
Template "top_menu" 800x480
   Button "Template_Button_3" at 3,3 size 45x34; TextOff 'Text'
      on Click: function_cf6f4242("GraphX_Slidein_Left", -1)
   Group "Group_2" at 3,3 size 45x34
   Group "Group_3" at 747,1 size 53x34
   GraphicView "Template_Graphic view_1" at 69,0 size 40x38; Picture "344330-200"
   Button "BtnBack" at 67,3 size 45x34; TextOff 'Text'
      on Click: function_efd93a16()
   GraphicView "Template_Graphic view_2" at 130,3 size 35x34; Picture "Artboard_43-512"
   Button "BtnHome" at 127,4 size 45x34; TextOff 'Text'
      on Click: ActivateScreen("Main", 0)
   IOField "Template_I/O field_2" at 638,2 size 46x16; FormatPattern 999; Unit  
   IOField "Template_I/O field_3" at 532,18 size 82x16; FormatPattern 999; Unit  
   TextField "Template_Text field_3" at 490,18 size 40x16; Text 'Errors:'
   IOField "Template_I/O field_1" at 614,18 size 70x16; FormatPattern 999; Unit  
   TextField "Template_Text field_1" at 619,19 size 27x16; Text 'Sim:'
   IOField "Template_I/O field_4" at 532,2 size 106x16; FormatPattern 999; Unit  
   TextField "Template_Text field_4" at 643,1 size 10x16; Text '/'
   TextField "Template_Text field_2" at 483,2 size 45x16; Text 'Alarms:'
   Button "Template_Button_2" at 531,1 size 154x34; TextOff 'Text'
   Switch "Template_Switch_1" at 684,1 size 64x34; CaptionText 'Switch'; TextOff 'Tags OFF'; TextOn 'Tags ON'
   Button "Template_Button_5" at 747,1 size 53x34; TextOff 'Text'
      on Click: function_cf6f4242("GraphX_Slidein_Right", -1)

screen "Main" 800x480, template "top_menu"
   ScreenModuleView "motorValveAnalogIcon_1" at 139,122 size 123x41; Guid_{11997190-91299} 'PT-01'; ScreenModuleType ""
      on Guid_{11997190-75677}: function_efd93a16("Analog1", 50, 50, -1, 0, 1)
   Group "Group" at 265,110 size 32x56
   Group "Group_1" at 56,180 size 42x20
   ScreenModuleView "analogInAndAlarmsIcon_1" at 533,124 size 73x71; Guid_{11997190-95263} 'MV-01'; ScreenModuleType ""
      on Guid_{11997190-75677}: function_efd93a16("Valve1", 30, 30, 1, -1, 1)
   ScreenModuleView "analogInAndAlarmsIcon_2" at 535,284 size 73x71; Guid_{11997190-95263} 'MV-02'; ScreenModuleType ""
      on Guid_{11997190-75677}: function_efd93a16("Valve2", 30, 30, 1, -1, 1)
   Group "Group_2" at 671,178 size 42x20
   Group "Group_3" at 668,342 size 42x20
   ScreenModuleView "motorValveAnalogIcon_2" at 144,282 size 123x41; Guid_{11997190-91299} 'TT-01'; ScreenModuleType ""
      on Guid_{11997190-75677}: function_efd93a16("Analog2", 50, 50, -1, 0, 1)
   TextField "Text field_1" at 269,115 size 24x23; Text 'PT'

PopupScreen "Analog1" 502x247
   ScreenModuleView "analogInAndAlarmsFP_1" at 1,1 size 500x244; ScreenModuleType ""
      Guid_{11997190-61144} <- "example_AI_PT44"
   Button "Button_1" at 429,9 size 57x36; TextOff 'X'
      on Click: function_efd93a16("Analog1", 30, 30, 0, -1, 1)

PopupScreen "Valve1" 502x247
   ScreenModuleView "motorValveFacplate_1" at 2,3 size 499x244; Guid_{11997190-89252} 'Valve 1'; ScreenModuleType ""
      on Guid_{11997190-86333}: function_efd93a16("Valve1", 50, 50, 0, -1, 1)
      Guid_{11997190-61144} <- "example_motorValveAnalog_DB_valve1_hmi"

screen "Alarms" 800x480, template "top_menu"
   AlarmView "Alarm view_1" at 8,42 size 789x432

PopupScreen "Valve2" 502x247
   ScreenModuleView "motorValveFacplate_1" at 2,3 size 499x244; Guid_{11997190-89252} 'Valve_2'; ScreenModuleType ""
      on Guid_{11997190-86333}: function_efd93a16("Valve2", 50, 50, 0, -1, 1)
      Guid_{11997190-61144} <- "example_motorValveAnalog_DB_valve2_hmi"

PopupScreen "Analog2" 502x247
   ScreenModuleView "analogInAndAlarmsFP_1" at 1,1 size 500x244; ScreenModuleType ""
      Guid_{11997190-61144} <- "example_AI_PT44"
   Button "Button_1" at 429,9 size 57x36; TextOff 'X'
      on Click: function_efd93a16("Analog2", 30, 30, 0, -1, 1)

screen "UserMangement" 800x480, template "top_menu"
   UserView "User view_1" at 7,46 size 782x425

screen "Diagnostics" 800x480, template "top_menu"
   SysDiagControl "System diagnostics view_1" at 3,40 size 792x436

screen "Test" 800x480, template "top_menu"
   PLCCodeViewer "PLC code view_1" at 35,84 size 543x266
   S7GraphOverview "GRAPH overview_1" at 159,383 size 424x72

screen "load_balanser" 800x480
   ScreenModuleView "load_balancer_faceplate_1" at 127,122 size 640x320; ScreenModuleType ""

VB script "VBFunction_1"
   'Tip:
   ' 1. Use the <CTRL+SPACE> or <CTRL+I> shortcut to open a list of all objects and functions
   ' 2. Write the code using the HMI Runtime object.
   '  Example: HmiRuntime.Screens("Screen_1").
   ' 3. Use the <CTRL+J> shortcut to create an object reference.
   'Write the code as of this position:
*)

(* ===== HMI "HMI_RT_1" =====
system functions are stored by id; their names below are inferred from use

ScreenModuleEditorView "AnalogInAndAlarmsIcon" 125x43
   Button "value_alarmH" at 104,17 size 16x12; TextOff 'H'
      on Click: SetTag("screen", 3)
      Visibility <- "aiUdt.alarmH.Q"
   Button "value_alarmL" at 104,26 size 16x12; TextOff 'L'
      on Click: SetTag("screen", 3)
      Visibility <- "aiUdt.alarmL.Q"
   Button "value_simulation" at 1,17 size 12x21; TextOff 'SIM'
      Visibility <- "aiUdt.ai.sim"
      Appearance <- "aiUdt.ai.sim"
   IOField "value_value" at 12,17 size 92x21; FormatPattern 99999.99
      ProcessValue <- "aiUdt.ai.Q"
      Appearance <- "aiUdt.ai.Error"
   Button "value_alarmLL" at 104,26 size 16x12; TextOff 'LL'
      on Click: SetTag("screen", 3)
      Visibility <- "aiUdt.alarmLL.Q"
   Button "value_alarmHH" at 104,17 size 16x12; TextOff 'HH'
      on Click: SetTag("screen", 3)
      Visibility <- "aiUdt.alarmHH.Q"
   Button "Button" at 0,1 size 123x40; TextOff 'Text'
   TextField "Text field_1" at 8,-1 size 91x20; Text 'TAG_TAG_TAG'
      Visibility <- "aiUdt.hmi.showTag"

VB script "unitIntervalChange"
   'Tip:
   ' 1. Use the <CTRL+SPACE> or <CTRL+I> shortcut to open a list of all objects and functions
   ' 2. Write the code using the HMI Runtime object. Example: HmiRuntime.Screens("Screen_1").
   ' 3. Use the <CTRL+J> shortcut to create an object reference.
*)

(* ===== HMI "HMI_RT_1" =====
system functions are stored by id; their names below are inferred from use

HMI tags "Default tag table"
   "screen" : Int, internal
   "unitIntervalPerCent" : Real, internal

ScreenModuleEditorView "analogInAndAlarmsFacplate" 500x244
   IOField "I/O field_13" at 228,60 size 66x30; FormatPattern 9999.99
      Visibility <- "screen"
      ProcessValue <- "aiUdt.ai.scaleMin"
   IOField "I/O field_14" at 228,98 size 66x30; FormatPattern 9999.99
      Visibility <- "screen"
      ProcessValue <- "aiUdt.ai.scaleMax"
   IOField "I/O field_15" at 228,140 size 66x30; FormatPattern 9999.99
      Visibility <- "screen"
   IOField "I/O field_16" at 228,178 size 66x30; FormatPattern 9999.99
      Visibility <- "screen"
   IOField "I/O field_17" at 71,59 size 77x30; FormatPattern 99999.99
      Visibility <- "screen"
      ProcessValue <- "aiUdt.ai.Q"
      ObjectEnable <- "aiUdt.ai.sim"
   TextField "Text field_8" at 157,64 size 65x20; Text 'Scale Min:'
      Visibility <- "screen"
   TextField "Text field_9" at 157,101 size 68x20; Text 'Scale Max:'
      Visibility <- "screen"
   TextField "Text field_10" at 157,144 size 46x20; Text 'Factor:'
      Visibility <- "screen"
   TextField "Text field_11" at 157,181 size 33x20; Text 'Bias:'
      Visibility <- "screen"
   TextField "Text field_12" at 7,65 size 42x20; Text 'Value:'
      Visibility <- "screen"
   IOField "I/O field_18" at 407,93 size 69x30; FormatPattern 999; Unit  %
      Visibility <- "screen"
      ProcessValue <- "aiUdt.ai.filterConst"
   TextField "Text field_14" at 308,98 size 73x20; Text 'Error Action'
      Visibility <- "screen"
   IOField "I/O field_19" at 413,58 size 66x30; FormatPattern 999999
      Visibility <- "screen"
      ProcessValue <- "aiUdt.ai.filterConst"
   TextField "Text field_15" at 310,65 size 66x20; Text 'FilterConst'
      Visibility <- "screen"
   TextField "Text field_17" at 6,98 size 55x20; Text 'Simulate'
      Visibility <- "screen"
      Appearance <- "aiUdt.ai.sim"
   TextField "Text field_29" at 307,125 size 78x36; Text 'Force inside scale:'
      Visibility <- "screen"
   IOField "I/O field_23" at 69,136 size 78x30; FormatPattern 999.9; Unit  %
      Visibility <- "screen"
      ProcessValue <- "aiUdt.ai.unitInterval"
   TextField "Text field_30" at 6,143 size 54x20; Text 'Raw val.'
      Visibility <- "screen"
   Button "BtnHelpFilterConst" at 383,61 size 26x24; TextOff '?'
      Visibility <- "screen"
   GraphicView "Graphic view_4" at 32,194 size 32x19; Picture "kisspng-computer-icons-cut-copy-and-paste-copying-clip-a-options-vector-5adbf59dcb7576.1022898415243647018334"
      Visibility <- "screen"
   GraphicView "Graphic view_5" at 83,192 size 24x27; Picture "kisspng-computer-icons-clipboard-cut-copy-and-paste-5ae0cc5c36eb73.140446591524681820225"
      Visibility <- "screen"
   Button "BtnScreenEmpty_7" at 31,188 size 40x31; TextOff 'Text'
      on Click: SetTag(N, 1)
      Visibility <- "screen"
   Button "BtnScreenEmpty_6" at 81,185 size 36x36; TextOff 'Text'
      on Click: SetTag("screen", 201)
      Visibility <- "screen"
   Switch "Switch_2" at 411,134 size 61x30; TextOn 'On'; CaptionText 'Switch'; TextOff 'Off'
      Appearance <- "aiUdt.ai.forceInsideScale"
      ProcessValue <- "aiUdt.ai.forceInsideScale"
      Visibility <- "screen"
   Switch "Switch_1" at 101,96 size 46x25; TextOn 'On'; CaptionText 'Switch'; TextOff 'Off'
      Appearance <- "aiUdt.ai.sim"
      ProcessValue <- "aiUdt.ai.sim"
      Visibility <- "screen"
   Button "BtnScreenEmpty" at 407,179 size 62x40; TextOff '?'
      on Click: SetTag("screen", 300)
      Visibility <- "screen"
   Polyline "Polyline_7" at 428,153 size 25x56
      Visibility <- "screen"
   Rectangle "Rectangle_1" at 98,119 size 75x47
      Visibility <- "screen"
   Polyline "Polyline_1" at 32,127 size 56x25
      Visibility <- "screen"
   TextField "Text field_18" at 23,109 size 47x22; Text 'Raw in'
      Visibility <- "screen"
   TextField "Text field_19" at 103,131 size 64x22; Text 'Run. avg'
      Visibility <- "screen"
   Polyline "Polyline_2" at 189,127 size 56x25
      Visibility <- "screen"
   Rectangle "Rectangle_2" at 253,121 size 73x42
      Visibility <- "screen"
   TextField "Text field_20" at 258,131 size 65x22; Text 'Err check'
      Visibility <- "screen"
   Polyline "Polyline_3" at 125,59 size 25x56
      Visibility <- "screen"
   TextField "Text field_21" at 50,68 size 80x22; Text 'Filter const.'
      Visibility <- "screen"
   Polyline "Polyline_4" at 344,122 size 56x25
      Visibility <- "screen"
   Rectangle "Rectangle_3" at 399,122 size 73x42
      Visibility <- "screen"
   TextField "Text field_22" at 408,131 size 48x22; Text 'Scaling'
      Visibility <- "screen"
   Polyline "Polyline_5" at 420,57 size 25x56
      Visibility <- "screen"
   TextField "Text field_23" at 339,69 size 75x22; Text 'Min & Max'
      Visibility <- "screen"
   Rectangle "Rectangle_4" at 344,197 size 73x42
      Visibility <- "screen"
   TextField "Text field_24" at 151,211 size 59x22; Text 'Simulate'
      Visibility <- "screen"
   Polyline "Polyline_6" at 280,211 size 56x25
      Visibility <- "screen"
   TextField "Text field_25" at 299,206 size 91x22; Text 'Factor & bias'
      Visibility <- "screen"
   Polyline "Polyline_8" at 424,211 size 56x25
      Visibility <- "screen"
   TextField "Text field_26" at 444,195 size 16x22; Text 'Q'
      Visibility <- "screen"
   Button "value_alarmHH" at 18,147 size 36x26; TextOff 'HH'
      on Click: SetTag("screen", 3)
      Visibility <- "screen"
      Appearance <- "aiUdt.alarmHH.Q"
   Button "value_alarmH" at 57,147 size 36x26; TextOff 'H'
      on Click: SetTag("screen", 3)
      Visibility <- "screen"
      Appearance <- "aiUdt.alarmH.Q"
   Button "value_alarmL" at 96,147 size 36x26; TextOff 'L'
      on Click: SetTag("screen", 3)
      Visibility <- "screen"
      Appearance <- "aiUdt.alarmL.Q"
   Button "value_alarmLL" at 135,147 size 36x26; TextOff 'LL'
      on Click: SetTag("screen", 3)
      Visibility <- "screen"
      Appearance <- "aiUdt.alarmLL.Q"
   Button "value_simulation" at 41,184 size 99x35; TextOff 'Simulation'
      Visibility <- "screen"
      Appearance <- "aiUdt.ai.sim"
   Bar "Bar" at 200,63 size 66x171; MinimumValue 0; MaximumValue 100
      MinimumValue <- "aiUdt.ai.scaleMin"
      ProcessValue <- "aiUdt.ai.Q"
      MaximumValue <- "aiUdt.ai.scaleMax"
      Visibility <- "screen"
   IOField "value_value" at 18,74 size 151x42; FormatPattern 99999999; Unit         
      Visibility <- "screen"
      ProcessValue <- "aiUdt.alarmHH.delay"
      Appearance <- "aiUdt.ai.Error"
   GraphicView "Graphic 123" at 33,9 size 40x37; Picture "123-512"
   GraphicView "Graphic gear" at 182,7 size 40x37; Picture "setting-512"
   GraphicView "Graphic alarm" at 109,6 size 40x37; Picture "UI_Glyph_09_-13-512"
   Button "BtnScreenValue" at 22,4 size 57x42; TextOff 'Text'
      on Click: SetTag("screen", 0)
   Button "BtnScreenAlarms" at 97,4 size 57x42; TextOff 'Text'
      on Click: SetTag("screen", 100)
   Button "BtnScreenSetup" at 174,4 size 57x42; TextOff 'Text'
      on Click: SetTag("screen", 200)
   Switch "Switch_10" at 131,197 size 46x27; TextOn 'On'; CaptionText 'Switch'; TextOff 'Off'
      Appearance <- "aiUdt.ai.forceInsideScale"
      Visibility <- "screen"
      ProcessValue <- "aiUdt.alarmLL.autoAck"
   IOField "I/O field_5" at 190,160 size 62x30; FormatPattern 9999.99
      Visibility <- "screen"
      ProcessValue <- "aiUdt.alarmL.lim"
   IOField "I/O field_1" at 190,84 size 62x30; FormatPattern 9999.99
      Visibility <- "screen"
      ProcessValue <- "aiUdt.alarmHH.lim"
   TextField "Text field_1" at 7,91 size 64x20; Text 'Alarm HH:'
      Visibility <- "screen"
   TextField "Text field_2" at 205,63 size 26x17; Text 'Limit'
      Visibility <- "screen"
   TextField "Text field_3" at 268,63 size 56x17; Text 'Delay [ms]'
      Visibility <- "screen"
   IOField "I/O field_2" at 265,84 size 53x30; FormatPattern 99999
      Visibility <- "screen"
      ProcessValue <- "aiUdt.alarmHH.delay"
   IOField "I/O field_3" at 190,121 size 62x30; FormatPattern 9999.99
      Visibility <- "screen"
      ProcessValue <- "aiUdt.alarmH.lim"
   TextField "Text field_4" at 7,125 size 56x20; Text 'Alarm H:'
      Visibility <- "screen"
   IOField "I/O field_4" at 265,121 size 53x30; FormatPattern 99999
      Visibility <- "screen"
      ProcessValue <- "aiUdt.alarmH.delay"
   TextField "Text field_5" at 7,165 size 54x20; Text 'Alarm L:'
      Visibility <- "screen"
   IOField "I/O field_6" at 265,160 size 53x30; FormatPattern 99999
      Visibility <- "screen"
      ProcessValue <- "aiUdt.alarmL.delay"
   IOField "I/O field_7" at 190,197 size 62x30; FormatPattern 9999.99
      Visibility <- "screen"
      ProcessValue <- "aiUdt.alarmLL.lim"
   TextField "Text field_6" at 7,201 size 60x20; Text 'Alarm LL:'
      Visibility <- "screen"
   IOField "I/O field_8" at 265,197 size 53x30; FormatPattern 99999
      Visibility <- "screen"
      ProcessValue <- "aiUdt.alarmLL.delay"
   IOField "I/O field_9" at 331,84 size 67x30; FormatPattern 9999.99
      Visibility <- "screen"
      ProcessValue <- "aiUdt.alarmHH.hyst"
   TextField "Text field_7" at 337,63 size 55x17; Text 'Hysteresis'
      Visibility <- "screen"
   IOField "I/O field_10" at 331,121 size 67x30; FormatPattern 9999.99
      Visibility <- "screen"
      ProcessValue <- "aiUdt.alarmH.hyst"
   IOField "I/O field_11" at 331,160 size 67x30; FormatPattern 9999.99
      Visibility <- "screen"
      ProcessValue <- "aiUdt.alarmL.hyst"
   IOField "I/O field_12" at 331,197 size 67x30; FormatPattern 9999.99
      Visibility <- "screen"
      ProcessValue <- "aiUdt.alarmLL.hyst"
   TextField "Text field_13" at 131,61 size 48x17; Text 'Auto Ack'
      Visibility <- "screen"
   Button "Button_11" at 419,85 size 53x63; TextOff 'Ack. all alarms'
      on Click: SetTag("aiUdt.alarmHH.ack", 1); SetTag("aiUdt.alarmH.ack", 1); SetTag("aiUdt.alarmL.ack", 1); SetTag("aiUdt.alarmLL.ack", 1)
      Visibility <- "screen"
   Switch "Switch_3" at 73,84 size 46x27; TextOn 'On'; CaptionText 'Switch'; TextOff 'Off'
      Appearance <- "aiUdt.ai.forceInsideScale"
      Visibility <- "screen"
      ProcessValue <- "aiUdt.alarmHH.enable"
   TextField "Text field_16" at 77,61 size 37x17; Text 'Enable'
      Visibility <- "screen"
   Switch "Switch_4" at 73,121 size 46x27; TextOn 'On'; CaptionText 'Switch'; TextOff 'Off'
      Appearance <- "aiUdt.ai.forceInsideScale"
      Visibility <- "screen"
      ProcessValue <- "aiUdt.alarmH.enable"
   Switch "Switch_5" at 73,160 size 46x27; TextOn 'On'; CaptionText 'Switch'; TextOff 'Off'
      Appearance <- "aiUdt.ai.forceInsideScale"
      Visibility <- "screen"
      ProcessValue <- "aiUdt.alarmL.enable"
   Switch "Switch_6" at 73,197 size 46x27; TextOn 'On'; CaptionText 'Switch'; TextOff 'Off'
      Appearance <- "aiUdt.ai.forceInsideScale"
      Visibility <- "screen"
      ProcessValue <- "aiUdt.alarmLL.enable"
   Switch "Switch_7" at 131,84 size 46x27; TextOn 'On'; CaptionText 'Switch'; TextOff 'Off'
      Appearance <- "aiUdt.ai.forceInsideScale"
      Visibility <- "screen"
      ProcessValue <- "aiUdt.alarmHH.autoAck"
   Switch "Switch_8" at 131,121 size 46x27; TextOn 'On'; CaptionText 'Switch'; TextOff 'Off'
      Appearance <- "aiUdt.ai.forceInsideScale"
      Visibility <- "screen"
      ProcessValue <- "aiUdt.alarmH.autoAck"
   Switch "Switch_9" at 131,160 size 46x27; TextOn 'On'; CaptionText 'Switch'; TextOff 'Off'
      Appearance <- "aiUdt.ai.forceInsideScale"
      Visibility <- "screen"
      ProcessValue <- "aiUdt.alarmL.autoAck"
   Rectangle "Rectangle_5" at 98,85 size 266x118
      Visibility <- "screen"
   Button "value_alarmHH_1" at 236,154 size 72x34; TextOff 'Cancel'
      on Click: SetTag("screen", 200)
      Appearance <- "aiUdt.alarmHH.Q"
      Visibility <- "screen"
   TextField "Text field_28" at 118,103 size 197x22; Text 'Paste all settings and alarms?'
      Visibility <- "screen"
   Button "value_alarmHH_2" at 132,154 size 72x34; TextOff 'Paste'
      on Click: SetTag(N, 1)
      Appearance <- "aiUdt.alarmHH.Q"
      Visibility <- "screen"
   TextField "Text field_27" at 67,125 size 49x22; Text 'Alarms'

VB script "unitIntervalChange"
   'Tip:
   ' 1. Use the <CTRL+SPACE> or <CTRL+I> shortcut to open a list of all objects and functions
   ' 2. Write the code using the HMI Runtime object. Example: HmiRuntime.Screens("Screen_1").
   ' 3. Use the <CTRL+J> shortcut to create an object reference.
   
   
   'SmartTags("unitIntervalPerCent") = SmartTags("Properties\aiUdt.ai.unitInterval") * 100;
*)

(* ===== HMI "HMI_RT_1" =====
system functions are stored by id; their names below are inferred from use

ScreenModuleEditorView "device_faceplate" 300x200
   TextField "Text field_2" at 5,10 size 130x20; Text 'Available:'
   TextField "Text field_3" at 8,36 size 130x20; Text 'In operation:'
   TextField "Text field_4" at 17,71 size 121x20; Text 'Operating time:'
   Button "Button_1" at 52,106 size 96x32; TextOff 'Force start'
      on Click: SetTag("PLC.Q", 1)
   Button "Button_2" at 175,106 size 96x32; TextOff 'Force stop'
      on Click: SetTag("PLC.Q", 0)
   IOField "I/O field_7" at 142,69 size 142x27; FormatPattern 9999999999; Unit  s
      ProcessValue <- "PLC.operation_time"
   Circle "Circle_1" at 141,12 size 17x17
      Appearance <- "PLC.available"
   Circle "Circle_2" at 141,37 size 18x18
      Appearance <- "PLC.in_operation"
   TextField "Text field_1" at 169,10 size 83x20; Text 'Started:'
   Circle "Circle_3" at 259,12 size 17x17
      Appearance <- "PLC.Q"
*)

(* ===== HMI "HMI_RT_1" =====
system functions are stored by id; their names below are inferred from use

HMI tags "Default tag table"
   "limit_above" : Bool, internal
   "limit_under" : Bool, internal
   "show_help" : Bool, internal

ScreenModuleEditorView "load_balancer_faceplate" 640x320
   Switch "Switch_1" at 549,82 size 71x24; TextOn 'ON'; CaptionText 'Switch'; TextOff 'OFF'
      ProcessValue <- "PLC.bypass"
      Appearance <- "PLC.bypass"
   TextField "Text field_1" at 358,83 size 183x20; Text 'Bypass load balancer:'
   IOField "I/O field_1" at 466,9 size 156x29; FormatPattern 9999
      ProcessValue <- "PLC.max_devices_same_time"
   TextField "Text field_2" at 231,13 size 229x20; Text 'Max oper. devices at same time:'
   TextField "Text field_3" at 159,44 size 229x20; Text 'Max diff. opeating time:'
   IOField "I/O field_2" at 466,40 size 156x29; FormatPattern 999999999; Unit  ms
      ProcessValue <- "PLC.max_diff_operating.sec"
   TextField "Text field_4" at 23,155 size 61x20; Text 'Limit:'
   TextField "Text field_5" at 23,188 size 61x20; Text 'Delay:'
   IOField "I/O field_3" at 90,146 size 114x29; FormatPattern 999; Unit  %
      ProcessValue <- "PLC.start.limit"
      Appearance <- "limit_above"
   IOField "I/O field_4" at 91,184 size 114x29; FormatPattern 999999; Unit  ms
      ProcessValue <- "PLC.start.delay"
   Button "Button_1" at 101,220 size 96x32; TextOff 'Force start'
      on Click: SetTag("PLC.start.force", 1)
   IOField "I/O field_5" at 211,145 size 114x29; FormatPattern 999; Unit  %
      ProcessValue <- "PLC.stop.limit"
      Appearance <- "limit_under"
   IOField "I/O field_6" at 211,182 size 114x29; FormatPattern 999999; Unit  ms
      ProcessValue <- "PLC.stop.delay"
   Button "Button_2" at 222,220 size 96x32; TextOff 'Force stop'
      on Click: SetTag("PLC.stop.force", 1)
   TextField "Text field_9" at 353,113 size 193x20; Text 'Devices total:'
   IOField "I/O field_7" at 549,112 size 71x22; FormatPattern 999
      ProcessValue <- "PLC.info.total"
   TextField "Text field_10" at 347,139 size 197x20; Text 'Devices in operation:'
   IOField "I/O field_8" at 549,138 size 71x22; FormatPattern 999
      ProcessValue <- "PLC.info.in_operation"
   TextField "Text field_11" at 348,163 size 198x20; Text 'Devices standby:'
   IOField "I/O field_9" at 549,164 size 71x22; FormatPattern 999
      ProcessValue <- "PLC.info.standby"
      Appearance <- "PLC.info.standby"
   TextField "Text field_6" at 12,82 size 314x20; Text 'Start and stop conditions'
   TextField "Text field_8" at 91,123 size 112x20; Text 'Start'
   TextField "Text field_12" at 214,123 size 109x20; Text 'Stop'
   TextField "Text field_13" at 20,18 size 199x20; Text 'Load balancer'
   TextField "Text field_14" at 224,78 size 105x20; Text 'Block input:'
   IOField "I/O field_10" at 260,98 size 71x22; FormatPattern 999; Unit  %
      ProcessValue <- "PLC.info.input"
   Switch "Switch_2" at 549,191 size 71x24; TextOn 'ON'; CaptionText 'Switch'; TextOff 'OFF'
      ProcessValue <- "PLC.bypass"
      Appearance <- "PLC.bypass"
   TextField "Text field_7" at 351,192 size 190x20; Text 'Enable boost start:'
   Switch "Switch_3" at 549,219 size 71x24; TextOn 'ON'; CaptionText 'Switch'; TextOff 'OFF'
      ProcessValue <- "PLC.bypass"
      Appearance <- "PLC.bypass"
   TextField "Text field_15" at 347,220 size 194x20; Text 'Boost start auto:'
   IOField "I/O field_11" at 547,247 size 73x29; FormatPattern 999
      Appearance <- "PLC.boostStart.auto"
   TextField "Text field_16" at 347,249 size 194x21; Text 'Boost start n devices:'
   Button "Button_3" at 549,280 size 73x28; TextOff 'Reset'
      on Click: SetTag("PLC.boostStart.reset", 1)
   TextField "Text field_17" at 347,277 size 194x33; Text 'Statistics for auto boost start:'
   Switch "Switch_4" at 391,43 size 70x24; TextOn 'ON'; CaptionText 'Switch'; TextOff 'OFF'
      ProcessValue <- "PLC.max_diff_operating.enable"
      Appearance <- "PLC.bypass"
   Button "Button_5" at 16,273 size 45x32; TextOff '?'
      on Click: SetTag("show_help", 1)
   Rectangle "Rectangle_4" at 45,43 size 567x249
      Visibility <- "show_help"
   TextField "Text field_19" at 63,61 size 536x216; Text '- If devices (eg. pumps) work in parallell, this function will start or stop devices to operate as the demand increase or decrease. - A devices will be added for operation, if #input is above a certain value for a ceratin time, eg above 90% for 50 seconds. Likewise a devices will be removed from operation if #input is bellow a certain value for a certain time, eg. 10% for 30 secunds. The limits and the times are adjustable. - It's the device with least operating time that will be added first, and the device with most operating hours will be removed from operation first. - #input will typically be the output of a pid-controller. - For vfd, there should be configured a ramp time to make a smooth transition when a device is added or removed for operation.'
      Visibility <- "show_help"
   Button "Button_4" at 546,57 size 54x40; TextOff 'X'
      on Click: SetTag("PLC.boostStart.reset", 1)
      Visibility <- "show_help"

VB script "input_change"
   SmartTags("limit_above") = SmartTags("PLC.info.input") > SmartTags("PLC.start.limit")
   
   SmartTags("limit_under") = SmartTags("PLC.info.input") < SmartTags("PLC.stop.limit")

VB script "test"
   'Tip:
   ' 1. Use the <CTRL+SPACE> or <CTRL+I> shortcut to open a list of all objects and functions
   ' 2. Write the code using the HMI Runtime object.
   '  Example: HmiRuntime.Screens("Screen_1").
   ' 3. Use the <CTRL+J> shortcut to create an object reference.
   'Write the code as of this position:
*)

(* ===== HMI "HMI_RT_1" =====

ScreenModuleEditorView "load_balancer_icon" 640x480
   TextField "Text field_10" at 9,50 size 108x20; Text 'Started:'
   IOField "I/O field_8" at 127,48 size 74x21; FormatPattern 999
   TextField "Text field_11" at 11,72 size 108x20; Text 'Standby:'
   IOField "I/O field_9" at 127,73 size 74x21; FormatPattern 999
      ProcessValue <- "PLC.info.standby"
   Button "Button_1" at 17,10 size 184x32; TextOff 'Load balancer'
*)

(* ===== HMI "HMI_RT_1" =====
system functions are stored by id; their names below are inferred from use

HMI tags "Default tag table"
   "screen" : Int, internal

text list "FailSafeAction": 0 'No action'; 1 'Open'; 2 'Close'

ScreenModuleEditorView "motorValveFacplate" 500x244
   Button "value_simulation" at 377,105 size 80x35; TextOff 'Manuel'
      on Activate: SetTag("udt.cmd.man", 1)
      Visibility <- "screen"
   IOField "value_value" at 79,97 size 69x27; FormatPattern 999; Unit  %
      Visibility <- "screen"
      ProcessValue <- "udt.io.in.pos"
   TextField "Text field_8" at 6,99 size 64x20; Text 'Feedback:'
      Visibility <- "screen"
   TextField "Text field_9" at 10,60 size 25x20; Text 'SP:'
      Visibility <- "screen"
   IOField "value_value_1" at 79,51 size 69x35; FormatPattern 999; Unit  %
      Visibility <- "screen"
      ProcessValue <- "udt.SP"
   Button "value_simulation_1" at 6,153 size 78x35; TextOff 'Open fully'
      on Activate: SetTag("udt.cmd.openFully", 1)
      Visibility <- "screen"
   Button "value_simulation_2" at 174,150 size 78x35; TextOff 'Close fully'
      on Activate: SetTag("udt.cmd.closeFully", 1)
      Visibility <- "screen"
   Button "value_simulation_3" at 5,197 size 78x35; TextOff 'Jog open'
      on Activate: SetTag("udt.cmd.jogOpen", 1)
      Visibility <- "screen"
   Button "value_simulation_4" at 174,194 size 78x35; TextOff 'Jog close'
      on Activate: SetTag("udt.cmd.jogClose", 1)
      Visibility <- "screen"
   Button "value_simulation_5" at 95,152 size 63x35; TextOff 'Stop'
      on Activate: SetTag("udt.cmd.stop", 1)
      Visibility <- "screen"
   Button "value_simulation_6" at 97,196 size 63x35; TextOff 'Reset'
      on Activate: SetTag("udt.cmd.reset", 1)
      Visibility <- "screen"
   TextField "Text field_10" at 257,49 size 73x22; Text 'Pos. error'
      Visibility <- "screen"
   TextField "Text field_11" at 329,49 size 63x22; Text 'Timeout'
      Visibility <- "screen"
   TextField "Text field_12" at 391,49 size 94x22; Text 'Quick timeout'
      Visibility <- "screen"
   Button "value_simulation_7" at 287,104 size 78x35; TextOff 'Auto'
      on Activate: SetTag("udt.cmd.man", 0)
      Visibility <- "screen"
   IOField "value_value_4" at 381,157 size 74x20; FormatPattern 999
      Visibility <- "screen"
   TextField "Text field_18" at 273,157 size 102x20; Text 'Operating hours:'
      Visibility <- "screen"
   IOField "value_value_3" at 381,181 size 74x20; FormatPattern 999
      Visibility <- "screen"
   TextField "Text field_19" at 273,181 size 80x20; Text 'Start counter'
      Visibility <- "screen"
   GraphicView "Graphic view_1" at 181,63 size 46x46; Picture "compter-Construction-crane-oil-gas-valve-fuel-sensor--512"
      Visibility <- "screen"
   TextField "Text field_1" at 257,70 size 62x22; Text 'Interllok'
      Visibility <- "screen"
   TextField "Text field_2" at 318,70 size 64x22; Text 'Fail safe'
      Visibility <- "screen"
   Bar "Bar" at 489,43 size 10x201; MinimumValue 0; MaximumValue 100
      ProcessValue <- "udt.io.in.pos"
      Appearance <- "udt.error.posError"
   Rectangle "Rectangle_5" at 98,85 size 266x118
      Visibility <- "screen"
   Button "value_alarmHH_1" at 236,154 size 72x34; TextOff 'Cancel'
      on Click: SetTag("screen", 200)
      Visibility <- "screen"
   TextField "Text field_28" at 118,103 size 197x22; Text 'Paste all settings and alarms?'
      Visibility <- "screen"
   Button "value_alarmHH_2" at 132,154 size 72x34; TextOff 'Paste'
      on Click: SetTag(N, 1)
      Visibility <- "screen"
   IOField "I/O field_20" at 176,63 size 77x22; FormatPattern 99999; Unit ms
      Visibility <- "screen"
      ProcessValue <- "udt.conf.longTimeout"
   TextField "Text field_27" at 67,65 size 52x20; Text 'Timeout'
      Visibility <- "screen"
   IOField "I/O field_21" at 173,127 size 77x22; FormatPattern s9999999999; Unit %
      Visibility <- "screen"
      ProcessValue <- "udt.conf.qucikTimeoutMinMovement"
   TextField "Text field_31" at 67,130 size 89x20; Text 'Min movement'
      Visibility <- "screen"
   IOField "I/O field_22" at 173,156 size 77x22; FormatPattern 99999; Unit ms
      Visibility <- "screen"
      ProcessValue <- "udt.conf.quickTimeoutIntervalCheaks"
   TextField "Text field_33" at 67,156 size 90x20; Text 'Interval checks'
      Visibility <- "screen"
   TextField "Text field_34" at 106,99 size 88x20; Text 'Quick timeout:'
      Visibility <- "screen"
   TextField "Text field_32" at 284,65 size 91x20; Text 'Fail safe action'
      Visibility <- "screen"
   TextField "Text field_37" at 316,100 size 64x20; Text 'Auto reset'
      Visibility <- "screen"
   SymbolicIOField "Symbolic I/O field_1" at 386,64 size 86x22; TextOn '1'; TextOff '0'; TextList "FailSafeAction"
      Visibility <- "screen"
      ProcessValue <- "udt.conf.feilSafeAction"
   Switch "Switch_11" at 207,96 size 43x25; TextOn 'On'; CaptionText 'Switch'; TextOff 'Off'
      Visibility <- "screen"
      ProcessValue <- "udt.conf.quickTimeoutEnable"
   Switch "Switch_12" at 428,94 size 43x25; TextOn 'On'; CaptionText 'Switch'; TextOff 'Off'
      Visibility <- "screen"
      ProcessValue <- "udt.conf.autoReset"
   Rectangle "Rectangle_9" at 67,94 size 187x90
      Visibility <- "screen"
   Button "closeWindow_5" at 70,97 size 28x28; TextOff 'i'
      Visibility <- "screen"
   Button "closeWindow_6" at 283,95 size 28x28; TextOff 'i'
      Visibility <- "screen"
   IOField "I/O field_24" at 368,150 size 111x22; FormatPattern 99999; Unit ms
      ProcessValue <- "udt.conf.gentleTimePauseBias"
      Visibility <- "screen"
   TextField "Text field_35" at 275,150 size 64x20; Text 'Pause min'
      Visibility <- "screen"
   IOField "I/O field_25" at 368,119 size 111x22; FormatPattern 99999; Unit ms
      Visibility <- "screen"
      ProcessValue <- "udt.conf.gentleTimeRun"
   TextField "Text field_36" at 275,87 size 32x20; Text 'Limit'
      Visibility <- "screen"
   TextField "Text field_38" at 56,91 size 115x20; Text 'Gentle open enable'
      Visibility <- "screen"
   TextField "Text field_39" at 55,122 size 116x20; Text 'Gentle close enable'
      Visibility <- "screen"
   IOField "I/O field_26" at 367,89 size 111x22; FormatPattern 99; Unit %
      Visibility <- "screen"
      ProcessValue <- "udt.conf.gentleActivteLowLimit"
   TextField "Text field_40" at 55,153 size 137x20; Text 'Gentle also on fail Safe'
      Visibility <- "screen"
   TextField "Text field_41" at 275,118 size 27x20; Text 'Run'
      Visibility <- "screen"
   Switch "Switch_13" at 211,87 size 43x25; TextOn 'On'; CaptionText 'Switch'; TextOff 'Off'
      Visibility <- "screen"
      ProcessValue <- "udt.conf.gentleOpenEnable"
   Switch "Switch_14" at 211,120 size 43x25; TextOn 'On'; CaptionText 'Switch'; TextOff 'Off'
      Visibility <- "screen"
      ProcessValue <- "udt.conf.gentleCloseEnable"
   Switch "Switch_15" at 211,153 size 43x25; TextOn 'On'; CaptionText 'Switch'; TextOff 'Off'
      Visibility <- "screen"
      ProcessValue <- "udt.conf.gentleAlsoOnFailSafe"
   Button "closeWindow_10" at 55,57 size 28x28; TextOff 'i'
      Visibility <- "screen"
   IOField "I/O field_1" at 368,182 size 111x22; FormatPattern 99999; Unit ms
      ProcessValue <- "udt.conf.gentleTimePauseDelta"
      Visibility <- "screen"
   TextField "Text field_3" at 275,182 size 71x20; Text 'Pause delta'
      Visibility <- "screen"
   IOField "I/O field_27" at 184,90 size 77x22; FormatPattern 99.9; Unit %
      Visibility <- "screen"
      ProcessValue <- "udt.conf.regModeMinOffset"
   TextField "Text field_42" at 121,60 size 68x20; Text 'Reg mode:'
      Visibility <- "screen"
   Switch "Switch_16" at 218,59 size 43x25; TextOn 'On'; CaptionText 'Switch'; TextOff 'Off'
      Visibility <- "screen"
      ProcessValue <- "udt.info.regMode"
   TextField "Text field_43" at 89,90 size 66x20; Text 'Min offset:'
      Visibility <- "screen"
   TextField "Text field_44" at 89,120 size 75x20; Text 'Time break:'
      Visibility <- "screen"
   IOField "I/O field_28" at 184,117 size 77x22; FormatPattern 99999; Unit ms
      Visibility <- "screen"
      ProcessValue <- "udt.conf.regModeTimeBreak"
   Rectangle "Rectangle_7" at 82,55 size 185x87
      Visibility <- "screen"
   TextField "Text field_45" at 310,62 size 124x20; Text 'No fully open switch:'
      Visibility <- "screen"
   Switch "Switch_17" at 437,61 size 43x25; TextOn 'On'; CaptionText 'Switch'; TextOff 'Off'
      Visibility <- "screen"
      ProcessValue <- "udt.conf.simFullyOpenWithPos"
   TextField "Text field_46" at 280,123 size 96x20; Text 'Limit fully open:'
      Visibility <- "screen"
   IOField "I/O field_29" at 402,122 size 77x22; FormatPattern 999.9; Unit %
      Visibility <- "screen"
      ProcessValue <- "udt.conf.fullyOpenPosLim"
   TextField "Text field_47" at 127,153 size 52x20; Text 'Pre stop'
      Visibility <- "screen"
   IOField "I/O field_30" at 185,153 size 77x22; FormatPattern 9.9; Unit %
      Visibility <- "screen"
      ProcessValue <- "udt.conf.preStop"
   TextField "Text field_48" at 280,94 size 132x20; Text 'No fully closed switch:'
      Visibility <- "screen"
   Switch "Switch_18" at 437,93 size 43x25; TextOn 'On'; CaptionText 'Switch'; TextOff 'Off'
      Visibility <- "screen"
      ProcessValue <- "udt.conf.simFullyClosedWithPos"
   TextField "Text field_49" at 280,152 size 104x20; Text 'Limit fully closed:'
      Visibility <- "screen"
   IOField "I/O field_31" at 402,151 size 77x22; FormatPattern 99.9; Unit %
      Visibility <- "screen"
      ProcessValue <- "udt.conf.fullyClosedPosLim"
   Rectangle "Rectangle_10" at 273,56 size 213x125
      Visibility <- "screen"
   Button "btnInfo_1" at 278,59 size 28x28; TextOff 'i'
      Visibility <- "screen"
   Button "btnInfo_2" at 89,151 size 28x28; TextOff 'i'
      Visibility <- "screen"
   Button "btnInfo_3" at 87,58 size 28x28; TextOff 'i'
      Visibility <- "screen"
   TextField "mmSim" at 280,25 size 32x18; Text 'Sim'
      Visibility <- "udt.sim.enable"
      Appearance <- "udt.sim.enable"
   GraphicView "Graphic valve" at 13,7 size 35x35; Picture "image2vector-6-512"
   GraphicView "Graphic gear" at 122,6 size 40x37; Picture "setting-512"
   TextField "Text field_20" at 311,25 size 39x18; Text 'Error'
      Visibility <- "screen"
   TextField "Text field_53" at 282,3 size 162x20; Text 'TAG_TAG_TAG_TAG_TAG'
   Button "closeWindow" at 441,1 size 57x42; TextOff 'X'
   GraphicView "Graphic gear_2" at 234,6 size 40x37; Picture "setting-512"
   GraphicView "Graphic gear_1" at 178,6 size 40x37; Picture "setting-512"
   GraphicView "Graphic view_2" at 69,7 size 36x33; Picture "kisspng-musical-theatre-computer-icons-vector-graphics-mas-amp-quot-5b6f175fcfee27.8210729615340071358517"
   TextField "Text_1" at 140,15 size 19x34; Text '1'
      Visibility <- "screen"
   TextField "Text_2" at 198,15 size 19x34; Text '2'
      Visibility <- "screen"
   TextField "Text_3" at 252,15 size 19x34; Text '3'
      Visibility <- "screen"
   TextField "mmSim_1" at 349,25 size 60x18; Text 'Prog sim'
      Visibility <- "udt.sim.simByPlc"
      Appearance <- "udt.sim.simByPlc"
   TextField "txtSimOnOff" at 8,76 size 118x20; Text 'Simulation of inputs'
      Visibility <- "screen"
   IOField "simVal" at 156,115 size 79x35; FormatPattern 999; Unit  %
      Visibility <- "screen"
      ProcessValue <- "udt.sim.pos"
   Switch "simOnOff" at 157,74 size 43x25; TextOn 'On'; CaptionText 'Switch'; TextOff 'Off'
      Visibility <- "screen"
      ProcessValue <- "udt.sim.enable"
   TextField "txtSimVal" at 6,124 size 139x20; Text 'Valve position feedback'
      Visibility <- "screen"
   TextField "txtSimDescrip" at 257,60 size 234x100; Text 'Simulation is useful during develpoing and comisning. It may be used in rare at cases on sites to disable interlooks. Simulation should only then be used at huge precoason. If misused it may create huge damge.'
      Visibility <- "screen"
   GraphicView "Graphic alarm" at 412,175 size 40x37; Picture "UI_Glyph_09_-13-512"
      Visibility <- "screen"
   Button "BtnScreenSetup_2" at 224,1 size 57x42; TextOff 'Text'
      on Click: SetTag("screen", 400)
   Button "BtnScreenSetup_1" at 168,1 size 57x42; TextOff 'Text'
      on Click: SetTag("screen", 300)
   Button "BtnScreenSetup" at 112,1 size 57x42; TextOff 'Text'
      on Click: SetTag("screen", 200)
   Button "BtnScreenSim" at 56,1 size 57x42; TextOff 'Text'
      on Click: SetTag("screen", 100)
   Button "BtnScreenValue" at 0,1 size 57x42; TextOff 'Text'
      on Click: SetTag("screen", 0)
   Rectangle "Background_1" at 35,27 size 386x147
      Visibility <- "screen"
   Button "closeWindow_7" at 41,33 size 374x138; TextOff 'Text'
      Visibility <- "screen"
   TextField "txtSettingsHelpGentle" at 74,59 size 299x68; Text 'Gentle open and close will force smal time breaks while the valve move under the specified limit. This may prevent huge pressure surge which may prevent a pipe to burst.'
      Visibility <- "screen"
   Rectangle "Background_2" at 43,35 size 386x147
      Visibility <- "screen"
   Button "closeWindow_8" at 49,41 size 374x138; TextOff 'Text'
      Visibility <- "screen"
   TextField "txtSettingsHelpQuciTimeout" at 82,67 size 343x84; Text 'Quick timeout At spesifed interval there will done checks to see if position move towards the setpoint. The minimum movment may also be spesifed. This give a quick error feedback compared to a normal timeout.'
      Visibility <- "screen"
   Rectangle "Background_3" at 51,43 size 386x147
      Visibility <- "screen"
   Button "closeWindow_9" at 57,49 size 374x138; TextOff 'Text'
      Visibility <- "screen"
   TextField "txtSettingsHelpQuciTimeout_1" at 90,75 size 315x52; Text 'Auto reset: A new setpint or anoter command will reset the valve, without the need to push the reset button first.'
      Visibility <- "screen"
   Rectangle "Background_4" at 59,51 size 386x147
      Visibility <- "screen"
   Button "closeWindow_12" at 65,57 size 374x138; TextOff 'Text'
      Visibility <- "screen"
   TextField "txtSettingsHelpQuciTimeout_2" at 98,83 size 63x20; Text 'Reg mode'
      Visibility <- "screen"
   Rectangle "Background_5" at 67,59 size 386x147
      Visibility <- "screen"
   Button "closeWindow_1" at 73,65 size 374x138; TextOff 'Text'
      Visibility <- "screen"
   TextField "txtSettingsHelpQuciTimeout_3" at 106,91 size 322x84; Text 'Pre stop: When the valve move towards the set point, it will stop about half a per centage before becouse it has some momentum. This features is disabled at almost closed and almost open position to avoid a dead lock situation.'
      Visibility <- "screen"
   Rectangle "Background_6" at 75,67 size 386x147
      Visibility <- "screen"
   Button "closeWindow_2" at 81,73 size 374x138; TextOff 'Text'
      Visibility <- "screen"
   TextField "txtSettingsHelpQuciTimeout_4" at 114,99 size 185x20; Text 'Fully open and fully close signal'
      Visibility <- "screen"

VB script "unitIntervalChange"
   'Tip:
   ' 1. Use the <CTRL+SPACE> or <CTRL+I> shortcut to open a list of all objects and functions
   ' 2. Write the code using the HMI Runtime object. Example: HmiRuntime.Screens("Screen_1").
   ' 3. Use the <CTRL+J> shortcut to create an object reference.
   
   
   SmartTags("unitIntervalPerCent") = SmartTags("aiUdt.ai.unitInterval") * 100;
*)

(* ===== HMI "HMI_RT_1" =====

HMI tags "Default tag table"
   "valveColor" : SInt, internal

ScreenModuleEditorView "motorValveIcon" 133x81
   Button "LabelOpening" at 43,32 size 23x8; TextOff 'Opening'
      Visibility <- "valveUdt.io.out.open"
   Button "LabelClosing" at 43,40 size 23x8; TextOff 'Closing'
      Visibility <- "valveUdt.io.out.close"
   Button "LabelFailSafe" at 3,38 size 23x8; TextOff 'Fail safe'
   Button "LabelFailSafe_1" at 9,63 size 30x8; TextOff 'Fail safe'
   Button "LabelFailSafe_3" at 39,63 size 30x8; TextOff 'Interlook'
   Button "Button" at 2,6 size 72x68; TextOff 'Text'
   Polygon "Polygon_1" at 9,46 size 44x17
      Appearance <- "valveColor"
   TextField "M" at 24,33 size 13x15; Text 'M'
   TextField "Text field_1" at 1,3 size 122x20; Text 'TAG_TAG_TAG_TAG'
   Button "LabelValueSimulation_1" at 1,17 size 41x10; TextOff 'SIM prog'
      Visibility <- "valveUdt.sim.simByPlc"
      Appearance <- "valveUdt.sim.simByPlc"
   Button "LabelValueSimulation" at 3,28 size 18x10; TextOff 'SIM'
      Visibility <- "valveUdt.sim.enable"
      Appearance <- "valveUdt.sim.enable"
   IOField "LabelPos" at 6,20 size 56x17; FormatPattern 999; Unit %
      ProcessValue <- "valveUdt.io.in.pos"

VB script "valveColor"
   'Error - red
   If SmartTags("valveUdt.io.in.posError")
   	Or SmartTags("valveUdt.error.timeout") 
   	Or SmartTags("valveUdt.error.posError") 
   Then	
   	SmartTags("valveColor") = 2 
   
   'Close - White
   ElseIf SmartTags("valveUdt.io.in.fullyClosed") Then
   	SmartTags("valveColor") = 3 
   
   'Open - Green
   ElseIf SmartTags("valveUdt.io.in.fullyOpen") Then
   	SmartTags("valveColor") = 5
   
   'Between - Yellow
   ElseIf SmartTags("valveUdt.io.in.fullyClosed")
   	And SmartTags("valveUdt.io.in.fullyOpen") 
   Then
   	SmartTags("valveColor") = 4 
   
   'Grey
   Else
   	SmartTags("valveColor") = 0 
   End	

VB script "a_info"
   'Tip:
   ' 1. Use the <CTRL+SPACE> or <CTRL+I> shortcut to open a list of all objects and functions
   ' 2. Write the code using the HMI Runtime object.
   '  Example: HmiRuntime.Screens("Screen_1").
   ' 3. Use the <CTRL+J> shortcut to create an object reference.
   'Write the code as of this position:
*)

(* ===== HMI "HMI_RT_1" =====

ScreenModuleEditorView "modbus_status" 500x300
   IOField "I/O field_1" at 168,76 size 213x22; FormatPattern 9999999
      ProcessValue <- "sbUdt.log.connected_time"
   TextField "Text field_1" at 18,78 size 146x20; Text 'Connected time:'
   IOField "I/O field_2" at 168,99 size 213x22; FormatPattern 9999999
      ProcessValue <- "sbUdt.log.disconnected_time"
   TextField "Text field_2" at 18,101 size 146x20; Text 'Disconnected time:'
   IOField "I/O field_3" at 168,122 size 115x22; FormatPattern 9999999999
      ProcessValue <- "sbUdt.log.done_cnt"
   Circle "Circle_2" at 169,53 size 19x19
      Appearance <- "sbUdt.out.error"
   TextField "Text field_3" at 18,125 size 146x20; Text 'Done cnt:'
   IOField "I/O field_4" at 168,145 size 115x22; FormatPattern 9999999999
      ProcessValue <- "sbUdt.log.error_exception_cnt"
   TextField "Text field_4" at 19,147 size 145x20; Text 'Exception cnt:'
   IOField "I/O field_5" at 168,168 size 115x22; FormatPattern 9999999999
      ProcessValue <- "sbUdt.out.error_comm"
   TextField "Text field_5" at 30,171 size 134x20; Text 'Comm. error cnt:'
   IOField "I/O field_6" at 168,191 size 115x22; FormatPattern FFFF
      ProcessValue <- "sbUdt.log.error_status"
   TextField "Text field_6" at 30,194 size 134x20; Text 'Error status:'
   TextField "Text field_7" at 15,30 size 147x20; Text 'Comm. error:'
   TextField "Text field_8" at 15,52 size 147x20; Text 'Error:'
   Circle "Circle_1" at 169,31 size 19x19
      Appearance <- "sbUdt.out.error_comm"
   IOField "I/O field_7" at 167,214 size 117x22; FormatPattern 999999
      ProcessValue <- "sbUdt.log.error_data_addr"
   TextField "Text field_9" at 24,215 size 141x20; Text 'Error data addr:'
   TextField "Text field_10" at 15,5 size 368x20; Text 'TAG_TAG_TAG_TAG_TAG_TAG_TAG_TAG_TAG_TAG'
*)

(* ===== HMI "HMI_RT_1" =====

ScreenModuleEditorView "modbus_conf" 400x150
   IOField "I/O field_8" at 168,79 size 117x22; FormatPattern 99999999
      ProcessValue <- "sbUdt.conf.max_comm_error"
   TextField "Text field_10" at 11,82 size 155x20; Text 'Conf. max.comm.err:'
   IOField "I/O field_9" at 168,55 size 117x22; FormatPattern 99999999
      ProcessValue <- "sbUdt.conf.exec_x_quries"
   TextField "Text field_11" at 11,58 size 155x20; Text 'Exec. n. queries:'
   Circle "Circle_3" at 170,33 size 19x19
      Appearance <- "sbUdt.conf.read_only"
   TextField "Text field_12" at 10,10 size 153x20; Text 'Disable:'
   TextField "Text field_13" at 10,32 size 153x20; Text 'Read only:'
   Circle "Circle_4" at 170,11 size 19x19
      Appearance <- "sbUdt.conf.disable"
*)